REGION Network 39
   RUNG wire#powerrail
      #"8#浊环热水泵引水电磁阀"(READY := wire#w1, HMI_OPEN :=, HMI_CLOSE :=, MA :=, AUTO :=, S :=, JT :=, "TIME" :=, OUT := "8#浊环热水泵引水电磁阀", TIME_OUT =>)
   END_RUNG
   RUNG wire#powerrail
      Contact( "8#浊环热水泵备妥" )
      Contact( "8#浊环热水电动蝶阀备妥" )
   END_RUNG wire#w1
   // the same network as SCL:
   #"8#浊环热水泵引水电磁阀"(READY := "8#浊环热水泵备妥" AND "8#浊环热水电动蝶阀备妥", OUT := "8#浊环热水泵引水电磁阀");   // "引水排气块"
END_REGION

REGION Network 40
   RUNG wire#powerrail
      #"8#浊环热水泵排气电磁阀"(READY := wire#w1, HMI_OPEN :=, HMI_CLOSE :=, MA :=, AUTO :=, S :=, JT :=, "TIME" :=, OUT := "8#浊环热水泵排气电磁阀", TIME_OUT =>)
   END_RUNG
   RUNG wire#powerrail
      Contact( "8#浊环热水泵备妥" )
      Contact( "8#浊环热水电动蝶阀备妥" )
   END_RUNG wire#w1
   // the same network as SCL:
   #"8#浊环热水泵排气电磁阀"(READY := "8#浊环热水泵备妥" AND "8#浊环热水电动蝶阀备妥", OUT := "8#浊环热水泵排气电磁阀");   // "引水排气块"
END_REGION

REGION Network 41
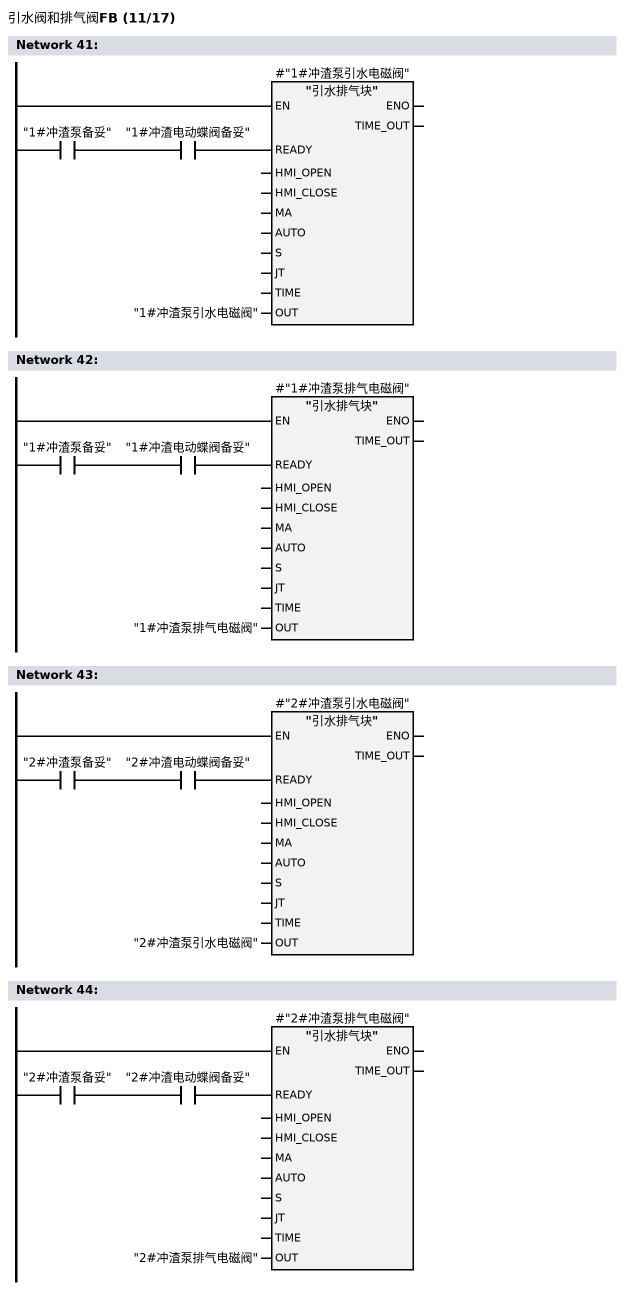
   RUNG wire#powerrail
      #"1#冲渣泵引水电磁阀"(READY := wire#w1, HMI_OPEN :=, HMI_CLOSE :=, MA :=, AUTO :=, S :=, JT :=, "TIME" :=, OUT := "1#冲渣泵引水电磁阀", TIME_OUT =>)
   END_RUNG
   RUNG wire#powerrail
      Contact( "1#冲渣泵备妥" )
      Contact( "1#冲渣电动蝶阀备妥" )
   END_RUNG wire#w1
   // the same network as SCL:
   #"1#冲渣泵引水电磁阀"(READY := "1#冲渣泵备妥" AND "1#冲渣电动蝶阀备妥", OUT := "1#冲渣泵引水电磁阀");   // "引水排气块"
END_REGION

REGION Network 42
   RUNG wire#powerrail
      #"1#冲渣泵排气电磁阀"(READY := wire#w1, HMI_OPEN :=, HMI_CLOSE :=, MA :=, AUTO :=, S :=, JT :=, "TIME" :=, OUT := "1#冲渣泵排气电磁阀", TIME_OUT =>)
   END_RUNG
   RUNG wire#powerrail
      Contact( "1#冲渣泵备妥" )
      Contact( "1#冲渣电动蝶阀备妥" )
   END_RUNG wire#w1
   // the same network as SCL:
   #"1#冲渣泵排气电磁阀"(READY := "1#冲渣泵备妥" AND "1#冲渣电动蝶阀备妥", OUT := "1#冲渣泵排气电磁阀");   // "引水排气块"
END_REGION

REGION Network 43
   RUNG wire#powerrail
      #"2#冲渣泵引水电磁阀"(READY := wire#w1, HMI_OPEN :=, HMI_CLOSE :=, MA :=, AUTO :=, S :=, JT :=, "TIME" :=, OUT := "2#冲渣泵引水电磁阀", TIME_OUT =>)
   END_RUNG
   RUNG wire#powerrail
      Contact( "2#冲渣泵备妥" )
      Contact( "2#冲渣电动蝶阀备妥" )
   END_RUNG wire#w1
   // the same network as SCL:
   #"2#冲渣泵引水电磁阀"(READY := "2#冲渣泵备妥" AND "2#冲渣电动蝶阀备妥", OUT := "2#冲渣泵引水电磁阀");   // "引水排气块"
END_REGION

REGION Network 44
   RUNG wire#powerrail
      #"2#冲渣泵排气电磁阀"(READY := wire#w1, HMI_OPEN :=, HMI_CLOSE :=, MA :=, AUTO :=, S :=, JT :=, "TIME" :=, OUT := "2#冲渣泵排气电磁阀", TIME_OUT =>)
   END_RUNG
   RUNG wire#powerrail
      Contact( "2#冲渣泵备妥" )
      Contact( "2#冲渣电动蝶阀备妥" )
   END_RUNG wire#w1
   // the same network as SCL:
   #"2#冲渣泵排气电磁阀"(READY := "2#冲渣泵备妥" AND "2#冲渣电动蝶阀备妥", OUT := "2#冲渣泵排气电磁阀");   // "引水排气块"
END_REGION

REGION Network 45
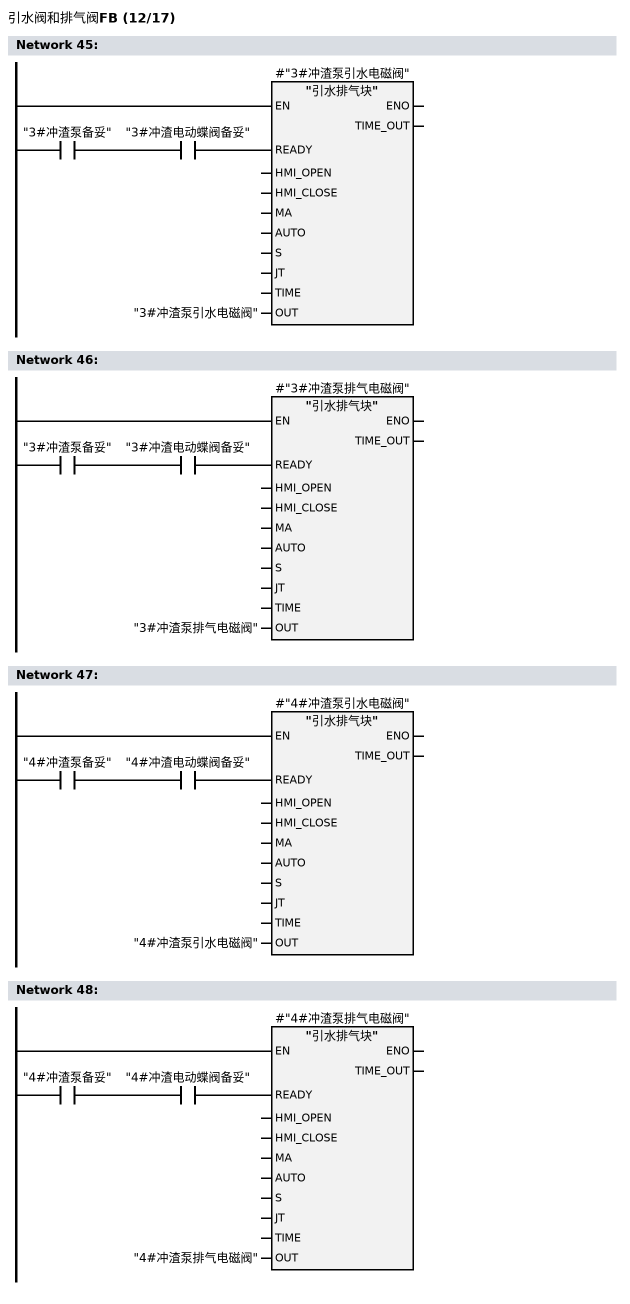
   RUNG wire#powerrail
      #"3#冲渣泵引水电磁阀"(READY := wire#w1, HMI_OPEN :=, HMI_CLOSE :=, MA :=, AUTO :=, S :=, JT :=, "TIME" :=, OUT := "3#冲渣泵引水电磁阀", TIME_OUT =>)
   END_RUNG
   RUNG wire#powerrail
      Contact( "3#冲渣泵备妥" )
      Contact( "3#冲渣电动蝶阀备妥" )
   END_RUNG wire#w1
   // the same network as SCL:
   #"3#冲渣泵引水电磁阀"(READY := "3#冲渣泵备妥" AND "3#冲渣电动蝶阀备妥", OUT := "3#冲渣泵引水电磁阀");   // "引水排气块"
END_REGION

REGION Network 46
   RUNG wire#powerrail
      #"3#冲渣泵排气电磁阀"(READY := wire#w1, HMI_OPEN :=, HMI_CLOSE :=, MA :=, AUTO :=, S :=, JT :=, "TIME" :=, OUT := "3#冲渣泵排气电磁阀", TIME_OUT =>)
   END_RUNG
   RUNG wire#powerrail
      Contact( "3#冲渣泵备妥" )
      Contact( "3#冲渣电动蝶阀备妥" )
   END_RUNG wire#w1
   // the same network as SCL:
   #"3#冲渣泵排气电磁阀"(READY := "3#冲渣泵备妥" AND "3#冲渣电动蝶阀备妥", OUT := "3#冲渣泵排气电磁阀");   // "引水排气块"
END_REGION

REGION Network 47
   RUNG wire#powerrail
      #"4#冲渣泵引水电磁阀"(READY := wire#w1, HMI_OPEN :=, HMI_CLOSE :=, MA :=, AUTO :=, S :=, JT :=, "TIME" :=, OUT := "4#冲渣泵引水电磁阀", TIME_OUT =>)
   END_RUNG
   RUNG wire#powerrail
      Contact( "4#冲渣泵备妥" )
      Contact( "4#冲渣电动蝶阀备妥" )
   END_RUNG wire#w1
   // the same network as SCL:
   #"4#冲渣泵引水电磁阀"(READY := "4#冲渣泵备妥" AND "4#冲渣电动蝶阀备妥", OUT := "4#冲渣泵引水电磁阀");   // "引水排气块"
END_REGION

REGION Network 48
   RUNG wire#powerrail
      #"4#冲渣泵排气电磁阀"(READY := wire#w1, HMI_OPEN :=, HMI_CLOSE :=, MA :=, AUTO :=, S :=, JT :=, "TIME" :=, OUT := "4#冲渣泵排气电磁阀", TIME_OUT =>)
   END_RUNG
   RUNG wire#powerrail
      Contact( "4#冲渣泵备妥" )
      Contact( "4#冲渣电动蝶阀备妥" )
   END_RUNG wire#w1
   // the same network as SCL:
   #"4#冲渣泵排气电磁阀"(READY := "4#冲渣泵备妥" AND "4#冲渣电动蝶阀备妥", OUT := "4#冲渣泵排气电磁阀");   // "引水排气块"
END_REGION

REGION Network 49
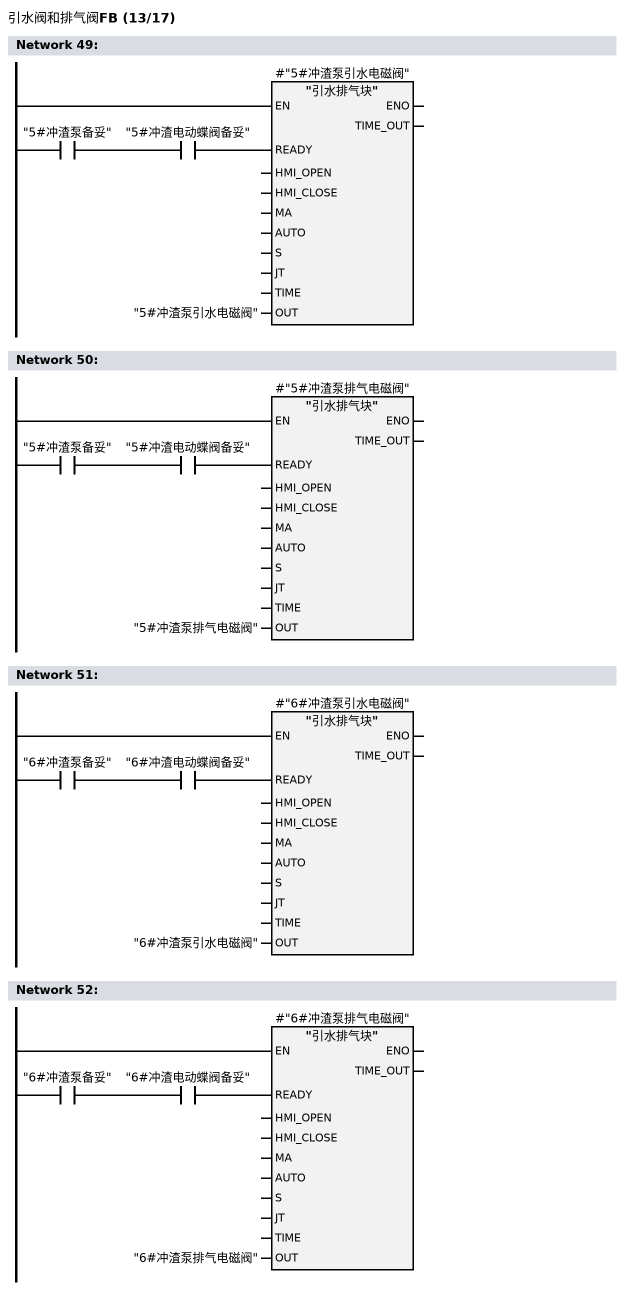
   RUNG wire#powerrail
      #"5#冲渣泵引水电磁阀"(READY := wire#w1, HMI_OPEN :=, HMI_CLOSE :=, MA :=, AUTO :=, S :=, JT :=, "TIME" :=, OUT := "5#冲渣泵引水电磁阀", TIME_OUT =>)
   END_RUNG
   RUNG wire#powerrail
      Contact( "5#冲渣泵备妥" )
      Contact( "5#冲渣电动蝶阀备妥" )
   END_RUNG wire#w1
   // the same network as SCL:
   #"5#冲渣泵引水电磁阀"(READY := "5#冲渣泵备妥" AND "5#冲渣电动蝶阀备妥", OUT := "5#冲渣泵引水电磁阀");   // "引水排气块"
END_REGION

REGION Network 50
   RUNG wire#powerrail
      #"5#冲渣泵排气电磁阀"(READY := wire#w1, HMI_OPEN :=, HMI_CLOSE :=, MA :=, AUTO :=, S :=, JT :=, "TIME" :=, OUT := "5#冲渣泵排气电磁阀", TIME_OUT =>)
   END_RUNG
   RUNG wire#powerrail
      Contact( "5#冲渣泵备妥" )
      Contact( "5#冲渣电动蝶阀备妥" )
   END_RUNG wire#w1
   // the same network as SCL:
   #"5#冲渣泵排气电磁阀"(READY := "5#冲渣泵备妥" AND "5#冲渣电动蝶阀备妥", OUT := "5#冲渣泵排气电磁阀");   // "引水排气块"
END_REGION

REGION Network 51
   RUNG wire#powerrail
      #"6#冲渣泵引水电磁阀"(READY := wire#w1, HMI_OPEN :=, HMI_CLOSE :=, MA :=, AUTO :=, S :=, JT :=, "TIME" :=, OUT := "6#冲渣泵引水电磁阀", TIME_OUT =>)
   END_RUNG
   RUNG wire#powerrail
      Contact( "6#冲渣泵备妥" )
      Contact( "6#冲渣电动蝶阀备妥" )
   END_RUNG wire#w1
   // the same network as SCL:
   #"6#冲渣泵引水电磁阀"(READY := "6#冲渣泵备妥" AND "6#冲渣电动蝶阀备妥", OUT := "6#冲渣泵引水电磁阀");   // "引水排气块"
END_REGION

REGION Network 52
   RUNG wire#powerrail
      #"6#冲渣泵排气电磁阀"(READY := wire#w1, HMI_OPEN :=, HMI_CLOSE :=, MA :=, AUTO :=, S :=, JT :=, "TIME" :=, OUT := "6#冲渣泵排气电磁阀", TIME_OUT =>)
   END_RUNG
   RUNG wire#powerrail
      Contact( "6#冲渣泵备妥" )
      Contact( "6#冲渣电动蝶阀备妥" )
   END_RUNG wire#w1
   // the same network as SCL:
   #"6#冲渣泵排气电磁阀"(READY := "6#冲渣泵备妥" AND "6#冲渣电动蝶阀备妥", OUT := "6#冲渣泵排气电磁阀");   // "引水排气块"
END_REGION

REGION Network 53
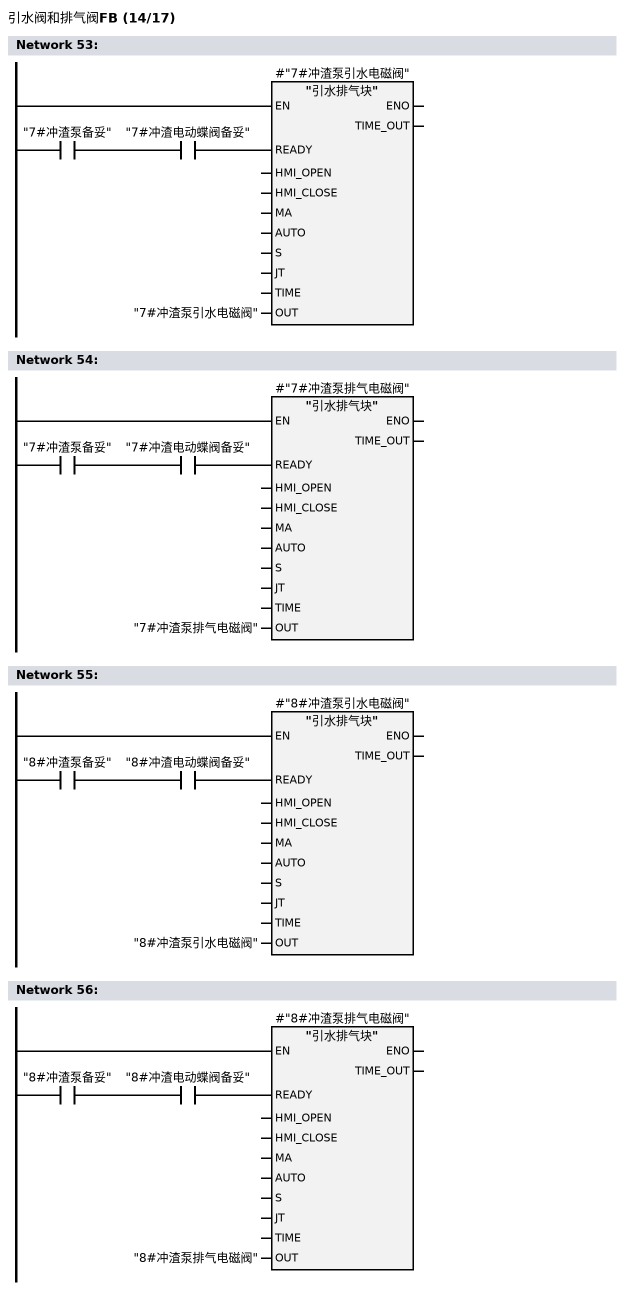
   RUNG wire#powerrail
      #"7#冲渣泵引水电磁阀"(READY := wire#w1, HMI_OPEN :=, HMI_CLOSE :=, MA :=, AUTO :=, S :=, JT :=, "TIME" :=, OUT := "7#冲渣泵引水电磁阀", TIME_OUT =>)
   END_RUNG
   RUNG wire#powerrail
      Contact( "7#冲渣泵备妥" )
      Contact( "7#冲渣电动蝶阀备妥" )
   END_RUNG wire#w1
   // the same network as SCL:
   #"7#冲渣泵引水电磁阀"(READY := "7#冲渣泵备妥" AND "7#冲渣电动蝶阀备妥", OUT := "7#冲渣泵引水电磁阀");   // "引水排气块"
END_REGION

REGION Network 54
   RUNG wire#powerrail
      #"7#冲渣泵排气电磁阀"(READY := wire#w1, HMI_OPEN :=, HMI_CLOSE :=, MA :=, AUTO :=, S :=, JT :=, "TIME" :=, OUT := "7#冲渣泵排气电磁阀", TIME_OUT =>)
   END_RUNG
   RUNG wire#powerrail
      Contact( "7#冲渣泵备妥" )
      Contact( "7#冲渣电动蝶阀备妥" )
   END_RUNG wire#w1
   // the same network as SCL:
   #"7#冲渣泵排气电磁阀"(READY := "7#冲渣泵备妥" AND "7#冲渣电动蝶阀备妥", OUT := "7#冲渣泵排气电磁阀");   // "引水排气块"
END_REGION

REGION Network 55
   RUNG wire#powerrail
      #"8#冲渣泵引水电磁阀"(READY := wire#w1, HMI_OPEN :=, HMI_CLOSE :=, MA :=, AUTO :=, S :=, JT :=, "TIME" :=, OUT := "8#冲渣泵引水电磁阀", TIME_OUT =>)
   END_RUNG
   RUNG wire#powerrail
      Contact( "8#冲渣泵备妥" )
      Contact( "8#冲渣电动蝶阀备妥" )
   END_RUNG wire#w1
   // the same network as SCL:
   #"8#冲渣泵引水电磁阀"(READY := "8#冲渣泵备妥" AND "8#冲渣电动蝶阀备妥", OUT := "8#冲渣泵引水电磁阀");   // "引水排气块"
END_REGION

REGION Network 56
   RUNG wire#powerrail
      #"8#冲渣泵排气电磁阀"(READY := wire#w1, HMI_OPEN :=, HMI_CLOSE :=, MA :=, AUTO :=, S :=, JT :=, "TIME" :=, OUT := "8#冲渣泵排气电磁阀", TIME_OUT =>)
   END_RUNG
   RUNG wire#powerrail
      Contact( "8#冲渣泵备妥" )
      Contact( "8#冲渣电动蝶阀备妥" )
   END_RUNG wire#w1
   // the same network as SCL:
   #"8#冲渣泵排气电磁阀"(READY := "8#冲渣泵备妥" AND "8#冲渣电动蝶阀备妥", OUT := "8#冲渣泵排气电磁阀");   // "引水排气块"
END_REGION

REGION Network 57
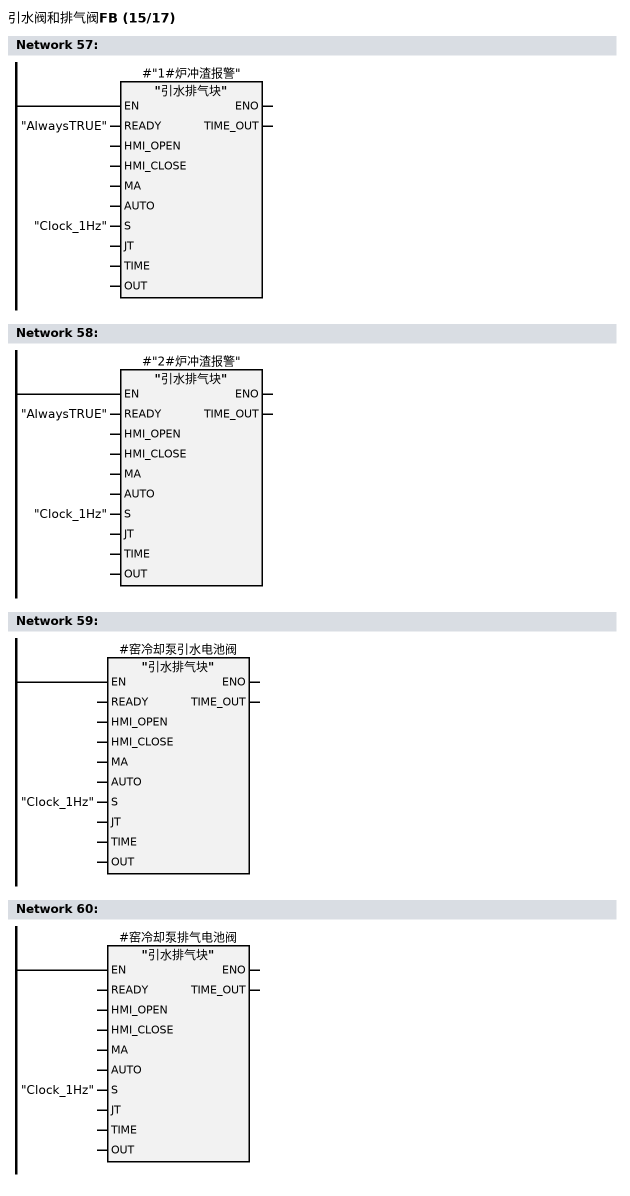
   RUNG wire#powerrail
      #"1#炉冲渣报警"(READY := "AlwaysTRUE", HMI_OPEN :=, HMI_CLOSE :=, MA :=, AUTO :=, S := "Clock_1Hz", JT :=, "TIME" :=, OUT :=, TIME_OUT =>)
   END_RUNG
   // the same network as SCL:
   #"1#炉冲渣报警"(READY := "AlwaysTRUE", S := "Clock_1Hz");   // "引水排气块"
END_REGION

REGION Network 58
   RUNG wire#powerrail
      #"2#炉冲渣报警"(READY := "AlwaysTRUE", HMI_OPEN :=, HMI_CLOSE :=, MA :=, AUTO :=, S := "Clock_1Hz", JT :=, "TIME" :=, OUT :=, TIME_OUT =>)
   END_RUNG
   // the same network as SCL:
   #"2#炉冲渣报警"(READY := "AlwaysTRUE", S := "Clock_1Hz");   // "引水排气块"
END_REGION

REGION Network 59
   RUNG wire#powerrail
      #窑冷却泵引水电池阀(READY :=, HMI_OPEN :=, HMI_CLOSE :=, MA :=, AUTO :=, S := "Clock_1Hz", JT :=, "TIME" :=, OUT :=, TIME_OUT =>)
   END_RUNG
   // the same network as SCL:
   #窑冷却泵引水电池阀(S := "Clock_1Hz");   // "引水排气块"
END_REGION

REGION Network 60
   RUNG wire#powerrail
      #窑冷却泵排气电池阀(READY :=, HMI_OPEN :=, HMI_CLOSE :=, MA :=, AUTO :=, S := "Clock_1Hz", JT :=, "TIME" :=, OUT :=, TIME_OUT =>)
   END_RUNG
   // the same network as SCL:
   #窑冷却泵排气电池阀(S := "Clock_1Hz");   // "引水排气块"
END_REGION

REGION Network 61
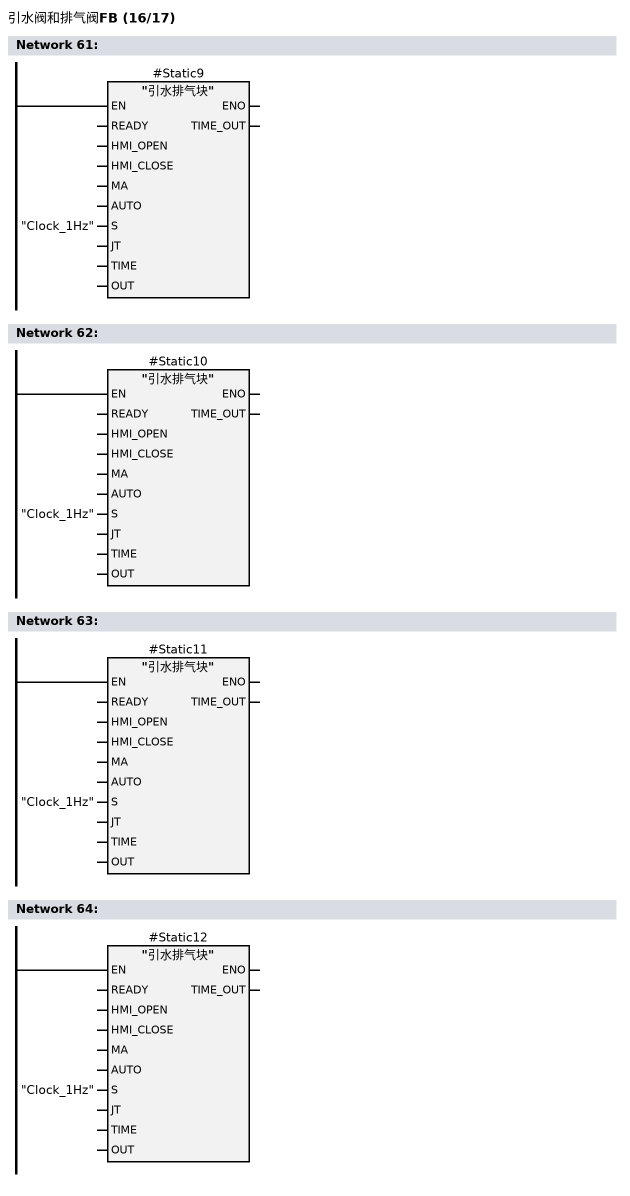
   RUNG wire#powerrail
      #Static9(READY :=, HMI_OPEN :=, HMI_CLOSE :=, MA :=, AUTO :=, S := "Clock_1Hz", JT :=, "TIME" :=, OUT :=, TIME_OUT =>)
   END_RUNG
   // the same network as SCL:
   #Static9(S := "Clock_1Hz");   // "引水排气块"
END_REGION

REGION Network 62
   RUNG wire#powerrail
      #Static10(READY :=, HMI_OPEN :=, HMI_CLOSE :=, MA :=, AUTO :=, S := "Clock_1Hz", JT :=, "TIME" :=, OUT :=, TIME_OUT =>)
   END_RUNG
   // the same network as SCL:
   #Static10(S := "Clock_1Hz");   // "引水排气块"
END_REGION

REGION Network 63
   RUNG wire#powerrail
      #Static11(READY :=, HMI_OPEN :=, HMI_CLOSE :=, MA :=, AUTO :=, S := "Clock_1Hz", JT :=, "TIME" :=, OUT :=, TIME_OUT =>)
   END_RUNG
   // the same network as SCL:
   #Static11(S := "Clock_1Hz");   // "引水排气块"
END_REGION

REGION Network 64
   RUNG wire#powerrail
      #Static12(READY :=, HMI_OPEN :=, HMI_CLOSE :=, MA :=, AUTO :=, S := "Clock_1Hz", JT :=, "TIME" :=, OUT :=, TIME_OUT =>)
   END_RUNG
   // the same network as SCL:
   #Static12(S := "Clock_1Hz");   // "引水排气块"
END_REGION

REGION Network 65
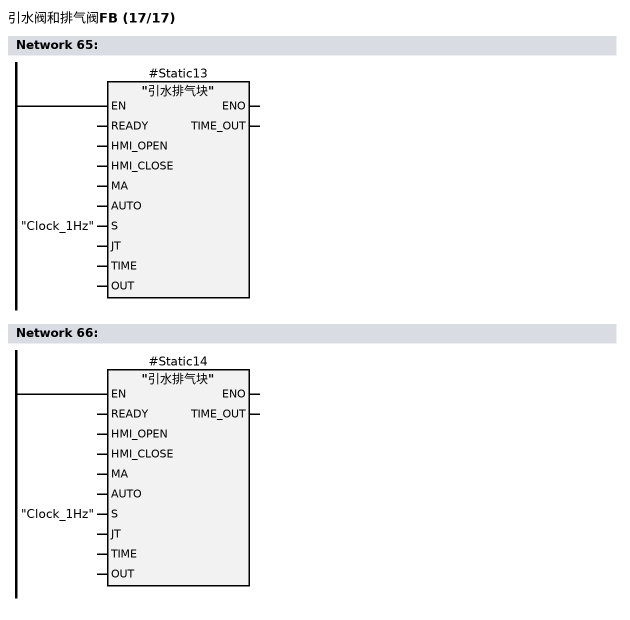
   RUNG wire#powerrail
      #Static13(READY :=, HMI_OPEN :=, HMI_CLOSE :=, MA :=, AUTO :=, S := "Clock_1Hz", JT :=, "TIME" :=, OUT :=, TIME_OUT =>)
   END_RUNG
   // the same network as SCL:
   #Static13(S := "Clock_1Hz");   // "引水排气块"
END_REGION

REGION Network 66
   RUNG wire#powerrail
      #Static14(READY :=, HMI_OPEN :=, HMI_CLOSE :=, MA :=, AUTO :=, S := "Clock_1Hz", JT :=, "TIME" :=, OUT :=, TIME_OUT =>)
   END_RUNG
   // the same network as SCL:
   #Static14(S := "Clock_1Hz");   // "引水排气块"
END_REGION
END_FUNCTION_BLOCK

FUNCTION_BLOCK "电机_泵FB"   // FB13, LAD
{ S7_Optimized_Access := 'FALSE' }
VERSION : 0.1
   VAR
      "1#冲渣泵驱动" : "电机_冷却塔风机";
      "2#冲渣泵驱动" : "电机_冷却塔风机";
      "3#冲渣泵驱动" : "电机_冷却塔风机";
      "4#冲渣泵驱动" : "电机_冷却塔风机";
      "5#冲渣泵驱动" : "电机_冷却塔风机";
      "6#冲渣泵驱动" : "电机_冷却塔风机";
      "7#冲渣泵驱动" : "电机_冷却塔风机";
      "8#冲渣泵驱动" : "电机_冷却塔风机";
      "1#浊环热水泵驱动" : "电机_冷却塔风机";
      "2#浊环热水泵驱动" : "电机_冷却塔风机";
      "3#浊环热水泵驱动" : "电机_冷却塔风机";
      "4#浊环热水泵驱动" : "电机_冷却塔风机";
      "5#浊环热水泵驱动" : "电机_冷却塔风机";
      "6#浊环热水泵驱动" : "电机_冷却塔风机";
      "7#浊环热水泵驱动" : "电机_冷却塔风机";
      "8#浊环热水泵驱动" : "电机_冷却塔风机";
      "1#炉体循环水泵驱动" : "电机_冷却塔风机";
      "2#炉体循环水泵驱动" : "电机_冷却塔风机";
      "3#炉体循环水泵驱动" : "电机_冷却塔风机";
      "1#电极循环水泵驱动" : "电机_冷却塔风机";
      "2#电极循环水泵驱动" : "电机_冷却塔风机";
      "3#电极循环水泵驱动" : "电机_冷却塔风机";
      "4#电极循环水泵驱动" : "电机_冷却塔风机";
      "1#净环热水泵驱动" : "电机_冷却塔风机";
      "2#净环热水泵驱动" : "电机_冷却塔风机";
      "3#净环热水泵驱动" : "电机_冷却塔风机";
      "4#净环热水泵驱动" : "电机_冷却塔风机";
      "5#净环热水泵驱动" : "电机_冷却塔风机";
      "1#柴油泵驱动" : "电机_冷却塔风机";
      "2#柴油泵驱动" : "电机_冷却塔风机";
      窑冷却泵驱动 : "电机_冷却塔风机";
      Static1 : "电机_冷却塔风机";
      Static2 : "电机_冷却塔风机";
      Static3 : "电机_冷却塔风机";
      Static4 : "电机_冷却塔风机";
      Static5 : "电机_冷却塔风机";
      Static6 : "电机_冷却塔风机";
      Static7 : "电机_冷却塔风机";
      Static8 : "电机_冷却塔风机";
      Static9 : "电机_冷却塔风机";
      Static10 : "电机_冷却塔风机";
      Static11 : "电机_冷却塔风机";
      Static12 : "电机_冷却塔风机";
      Static13 : "电机_冷却塔风机";
      Static14 : "电机_冷却塔风机";
      Static15 : "电机_冷却塔风机";
      Static16 : "电机_冷却塔风机";
      Static17 : "电机_冷却塔风机";
      Static18 : "电机_冷却塔风机";
      Static19 : "电机_冷却塔风机";
      Static20 : "电机_冷却塔风机";
      Static21 : "电机_冷却塔风机";
      Static22 : "电机_冷却塔风机";
      Static23 : "电机_冷却塔风机";
      Static24 : "电机_冷却塔风机";
      Static25 : "电机_冷却塔风机";
      Static26 : "电机_冷却塔风机";
      Static27 : "电机_冷却塔风机";
      Static28 : "电机_冷却塔风机";
      Static29 : "电机_冷却塔风机";
      Static30 : "电机_冷却塔风机";
      Static31 : "电机_冷却塔风机";
      Static32 : "电机_冷却塔风机";
      Static33 : "电机_冷却塔风机";
      Static34 : "电机_冷却塔风机";
      Static35 : "电机_冷却塔风机";
      Static36 : "电机_冷却塔风机";
      Static37 : "电机_冷却塔风机";
      Static38 : "电机_冷却塔风机";
      Static39 : "电机_冷却塔风机";
      Static40 : "电机_冷却塔风机";
      Static41 : "电机_冷却塔风机";
      Static42 : "电机_冷却塔风机";
      Static43 : "电机_冷却塔风机";
      Static44 : "电机_冷却塔风机";
      Static45 : "电机_冷却塔风机";
      Static46 : "电机_冷却塔风机";
      Static47 : "电机_冷却塔风机";
      Static48 : "电机_冷却塔风机";
      Static49 : "电机_冷却塔风机";
   END_VAR
BEGIN

REGION Network 1
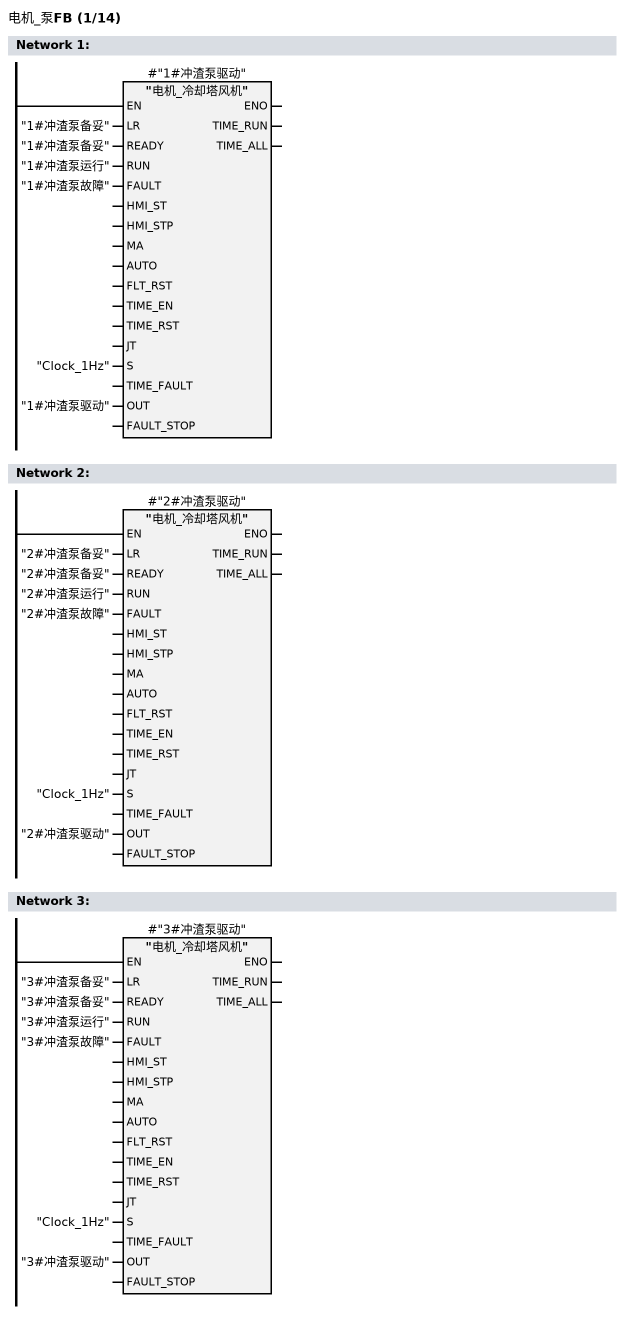
   RUNG wire#powerrail
      #"1#冲渣泵驱动"(LR := "1#冲渣泵备妥", READY := "1#冲渣泵备妥", RUN := "1#冲渣泵运行", FAULT := "1#冲渣泵故障", HMI_ST :=, HMI_STP :=, MA :=, AUTO :=, FLT_RST :=, TIME_EN :=, TIME_RST :=, JT :=, S := "Clock_1Hz", TIME_FAULT :=, OUT := "1#冲渣泵驱动", FAULT_STOP :=, TIME_RUN =>, TIME_ALL =>)
   END_RUNG
   // the same network as SCL:
   #"1#冲渣泵驱动"(LR := "1#冲渣泵备妥",   // "电机_冷却塔风机"
              READY := "1#冲渣泵备妥",
              RUN := "1#冲渣泵运行",
              FAULT := "1#冲渣泵故障",
              S := "Clock_1Hz",
              OUT := "1#冲渣泵驱动");
END_REGION

REGION Network 2
   RUNG wire#powerrail
      #"2#冲渣泵驱动"(LR := "2#冲渣泵备妥", READY := "2#冲渣泵备妥", RUN := "2#冲渣泵运行", FAULT := "2#冲渣泵故障", HMI_ST :=, HMI_STP :=, MA :=, AUTO :=, FLT_RST :=, TIME_EN :=, TIME_RST :=, JT :=, S := "Clock_1Hz", TIME_FAULT :=, OUT := "2#冲渣泵驱动", FAULT_STOP :=, TIME_RUN =>, TIME_ALL =>)
   END_RUNG
   // the same network as SCL:
   #"2#冲渣泵驱动"(LR := "2#冲渣泵备妥",   // "电机_冷却塔风机"
              READY := "2#冲渣泵备妥",
              RUN := "2#冲渣泵运行",
              FAULT := "2#冲渣泵故障",
              S := "Clock_1Hz",
              OUT := "2#冲渣泵驱动");
END_REGION

REGION Network 3
   RUNG wire#powerrail
      #"3#冲渣泵驱动"(LR := "3#冲渣泵备妥", READY := "3#冲渣泵备妥", RUN := "3#冲渣泵运行", FAULT := "3#冲渣泵故障", HMI_ST :=, HMI_STP :=, MA :=, AUTO :=, FLT_RST :=, TIME_EN :=, TIME_RST :=, JT :=, S := "Clock_1Hz", TIME_FAULT :=, OUT := "3#冲渣泵驱动", FAULT_STOP :=, TIME_RUN =>, TIME_ALL =>)
   END_RUNG
   // the same network as SCL:
   #"3#冲渣泵驱动"(LR := "3#冲渣泵备妥",   // "电机_冷却塔风机"
              READY := "3#冲渣泵备妥",
              RUN := "3#冲渣泵运行",
              FAULT := "3#冲渣泵故障",
              S := "Clock_1Hz",
              OUT := "3#冲渣泵驱动");
END_REGION

REGION Network 4
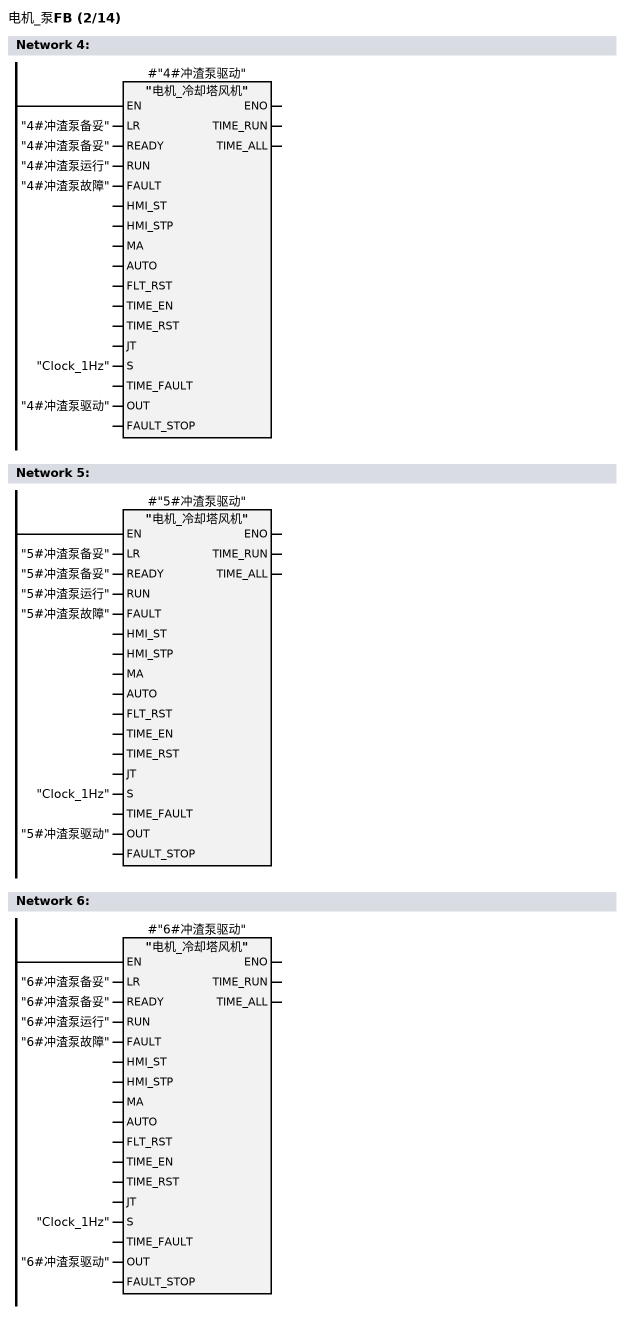
   RUNG wire#powerrail
      #"4#冲渣泵驱动"(LR := "4#冲渣泵备妥", READY := "4#冲渣泵备妥", RUN := "4#冲渣泵运行", FAULT := "4#冲渣泵故障", HMI_ST :=, HMI_STP :=, MA :=, AUTO :=, FLT_RST :=, TIME_EN :=, TIME_RST :=, JT :=, S := "Clock_1Hz", TIME_FAULT :=, OUT := "4#冲渣泵驱动", FAULT_STOP :=, TIME_RUN =>, TIME_ALL =>)
   END_RUNG
   // the same network as SCL:
   #"4#冲渣泵驱动"(LR := "4#冲渣泵备妥",   // "电机_冷却塔风机"
              READY := "4#冲渣泵备妥",
              RUN := "4#冲渣泵运行",
              FAULT := "4#冲渣泵故障",
              S := "Clock_1Hz",
              OUT := "4#冲渣泵驱动");
END_REGION

REGION Network 5
   RUNG wire#powerrail
      #"5#冲渣泵驱动"(LR := "5#冲渣泵备妥", READY := "5#冲渣泵备妥", RUN := "5#冲渣泵运行", FAULT := "5#冲渣泵故障", HMI_ST :=, HMI_STP :=, MA :=, AUTO :=, FLT_RST :=, TIME_EN :=, TIME_RST :=, JT :=, S := "Clock_1Hz", TIME_FAULT :=, OUT := "5#冲渣泵驱动", FAULT_STOP :=, TIME_RUN =>, TIME_ALL =>)
   END_RUNG
   // the same network as SCL:
   #"5#冲渣泵驱动"(LR := "5#冲渣泵备妥",   // "电机_冷却塔风机"
              READY := "5#冲渣泵备妥",
              RUN := "5#冲渣泵运行",
              FAULT := "5#冲渣泵故障",
              S := "Clock_1Hz",
              OUT := "5#冲渣泵驱动");
END_REGION

REGION Network 6
   RUNG wire#powerrail
      #"6#冲渣泵驱动"(LR := "6#冲渣泵备妥", READY := "6#冲渣泵备妥", RUN := "6#冲渣泵运行", FAULT := "6#冲渣泵故障", HMI_ST :=, HMI_STP :=, MA :=, AUTO :=, FLT_RST :=, TIME_EN :=, TIME_RST :=, JT :=, S := "Clock_1Hz", TIME_FAULT :=, OUT := "6#冲渣泵驱动", FAULT_STOP :=, TIME_RUN =>, TIME_ALL =>)
   END_RUNG
   // the same network as SCL:
   #"6#冲渣泵驱动"(LR := "6#冲渣泵备妥",   // "电机_冷却塔风机"
              READY := "6#冲渣泵备妥",
              RUN := "6#冲渣泵运行",
              FAULT := "6#冲渣泵故障",
              S := "Clock_1Hz",
              OUT := "6#冲渣泵驱动");
END_REGION

REGION Network 7
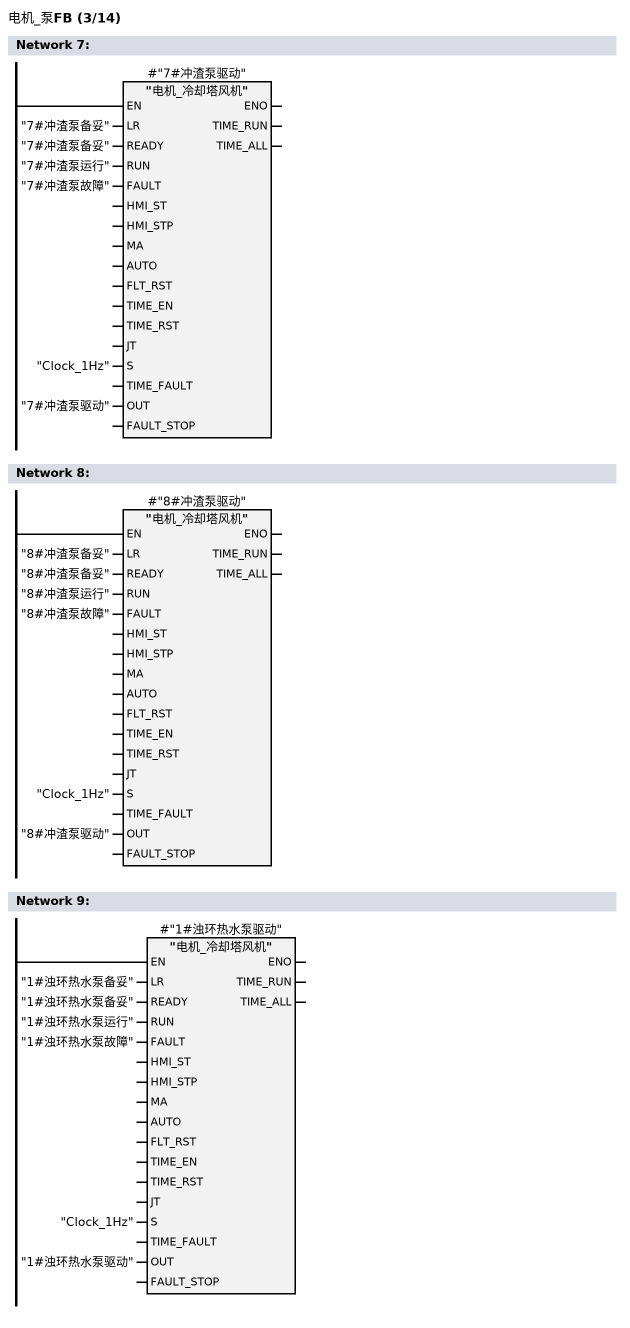
   RUNG wire#powerrail
      #"7#冲渣泵驱动"(LR := "7#冲渣泵备妥", READY := "7#冲渣泵备妥", RUN := "7#冲渣泵运行", FAULT := "7#冲渣泵故障", HMI_ST :=, HMI_STP :=, MA :=, AUTO :=, FLT_RST :=, TIME_EN :=, TIME_RST :=, JT :=, S := "Clock_1Hz", TIME_FAULT :=, OUT := "7#冲渣泵驱动", FAULT_STOP :=, TIME_RUN =>, TIME_ALL =>)
   END_RUNG
   // the same network as SCL:
   #"7#冲渣泵驱动"(LR := "7#冲渣泵备妥",   // "电机_冷却塔风机"
              READY := "7#冲渣泵备妥",
              RUN := "7#冲渣泵运行",
              FAULT := "7#冲渣泵故障",
              S := "Clock_1Hz",
              OUT := "7#冲渣泵驱动");
END_REGION

REGION Network 8
   RUNG wire#powerrail
      #"8#冲渣泵驱动"(LR := "8#冲渣泵备妥", READY := "8#冲渣泵备妥", RUN := "8#冲渣泵运行", FAULT := "8#冲渣泵故障", HMI_ST :=, HMI_STP :=, MA :=, AUTO :=, FLT_RST :=, TIME_EN :=, TIME_RST :=, JT :=, S := "Clock_1Hz", TIME_FAULT :=, OUT := "8#冲渣泵驱动", FAULT_STOP :=, TIME_RUN =>, TIME_ALL =>)
   END_RUNG
   // the same network as SCL:
   #"8#冲渣泵驱动"(LR := "8#冲渣泵备妥",   // "电机_冷却塔风机"
              READY := "8#冲渣泵备妥",
              RUN := "8#冲渣泵运行",
              FAULT := "8#冲渣泵故障",
              S := "Clock_1Hz",
              OUT := "8#冲渣泵驱动");
END_REGION

REGION Network 9
   RUNG wire#powerrail
      #"1#浊环热水泵驱动"(LR := "1#浊环热水泵备妥", READY := "1#浊环热水泵备妥", RUN := "1#浊环热水泵运行", FAULT := "1#浊环热水泵故障", HMI_ST :=, HMI_STP :=, MA :=, AUTO :=, FLT_RST :=, TIME_EN :=, TIME_RST :=, JT :=, S := "Clock_1Hz", TIME_FAULT :=, OUT := "1#浊环热水泵驱动", FAULT_STOP :=, TIME_RUN =>, TIME_ALL =>)
   END_RUNG
   // the same network as SCL:
   #"1#浊环热水泵驱动"(LR := "1#浊环热水泵备妥",   // "电机_冷却塔风机"
                READY := "1#浊环热水泵备妥",
                RUN := "1#浊环热水泵运行",
                FAULT := "1#浊环热水泵故障",
                S := "Clock_1Hz",
                OUT := "1#浊环热水泵驱动");
END_REGION

REGION Network 10
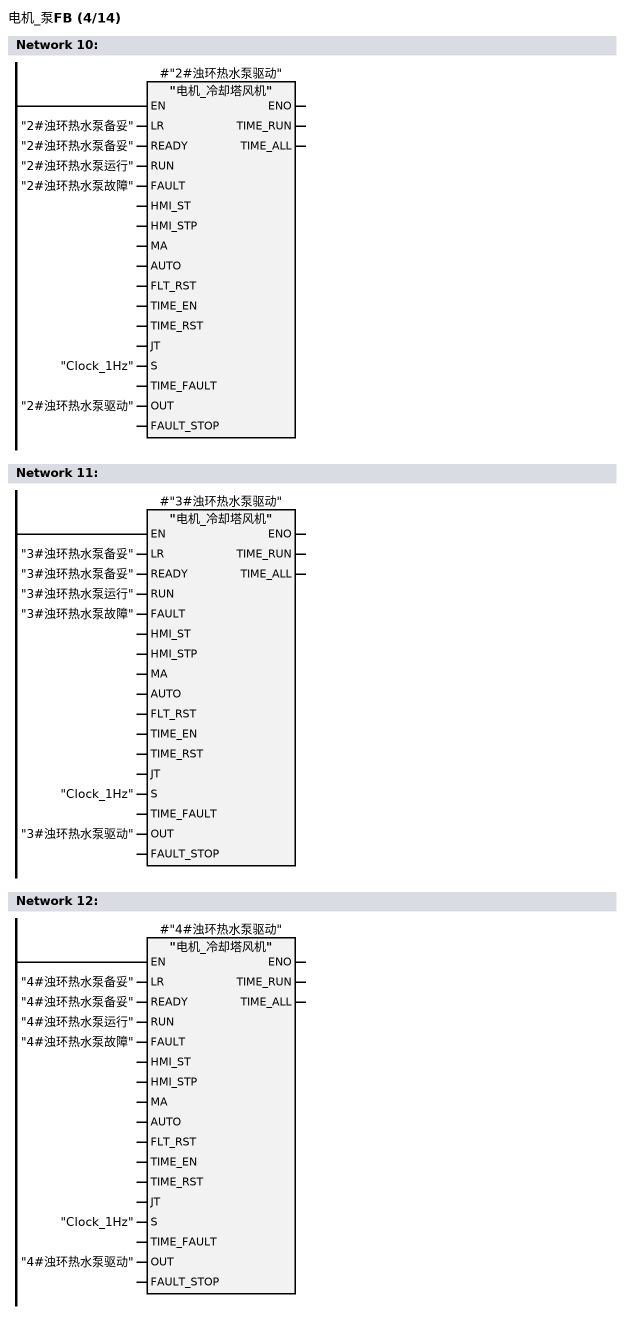
   RUNG wire#powerrail
      #"2#浊环热水泵驱动"(LR := "2#浊环热水泵备妥", READY := "2#浊环热水泵备妥", RUN := "2#浊环热水泵运行", FAULT := "2#浊环热水泵故障", HMI_ST :=, HMI_STP :=, MA :=, AUTO :=, FLT_RST :=, TIME_EN :=, TIME_RST :=, JT :=, S := "Clock_1Hz", TIME_FAULT :=, OUT := "2#浊环热水泵驱动", FAULT_STOP :=, TIME_RUN =>, TIME_ALL =>)
   END_RUNG
   // the same network as SCL:
   #"2#浊环热水泵驱动"(LR := "2#浊环热水泵备妥",   // "电机_冷却塔风机"
                READY := "2#浊环热水泵备妥",
                RUN := "2#浊环热水泵运行",
                FAULT := "2#浊环热水泵故障",
                S := "Clock_1Hz",
                OUT := "2#浊环热水泵驱动");
END_REGION

REGION Network 11
   RUNG wire#powerrail
      #"3#浊环热水泵驱动"(LR := "3#浊环热水泵备妥", READY := "3#浊环热水泵备妥", RUN := "3#浊环热水泵运行", FAULT := "3#浊环热水泵故障", HMI_ST :=, HMI_STP :=, MA :=, AUTO :=, FLT_RST :=, TIME_EN :=, TIME_RST :=, JT :=, S := "Clock_1Hz", TIME_FAULT :=, OUT := "3#浊环热水泵驱动", FAULT_STOP :=, TIME_RUN =>, TIME_ALL =>)
   END_RUNG
   // the same network as SCL:
   #"3#浊环热水泵驱动"(LR := "3#浊环热水泵备妥",   // "电机_冷却塔风机"
                READY := "3#浊环热水泵备妥",
                RUN := "3#浊环热水泵运行",
                FAULT := "3#浊环热水泵故障",
                S := "Clock_1Hz",
                OUT := "3#浊环热水泵驱动");
END_REGION

REGION Network 12
   RUNG wire#powerrail
      #"4#浊环热水泵驱动"(LR := "4#浊环热水泵备妥", READY := "4#浊环热水泵备妥", RUN := "4#浊环热水泵运行", FAULT := "4#浊环热水泵故障", HMI_ST :=, HMI_STP :=, MA :=, AUTO :=, FLT_RST :=, TIME_EN :=, TIME_RST :=, JT :=, S := "Clock_1Hz", TIME_FAULT :=, OUT := "4#浊环热水泵驱动", FAULT_STOP :=, TIME_RUN =>, TIME_ALL =>)
   END_RUNG
   // the same network as SCL:
   #"4#浊环热水泵驱动"(LR := "4#浊环热水泵备妥",   // "电机_冷却塔风机"
                READY := "4#浊环热水泵备妥",
                RUN := "4#浊环热水泵运行",
                FAULT := "4#浊环热水泵故障",
                S := "Clock_1Hz",
                OUT := "4#浊环热水泵驱动");
END_REGION

REGION Network 13
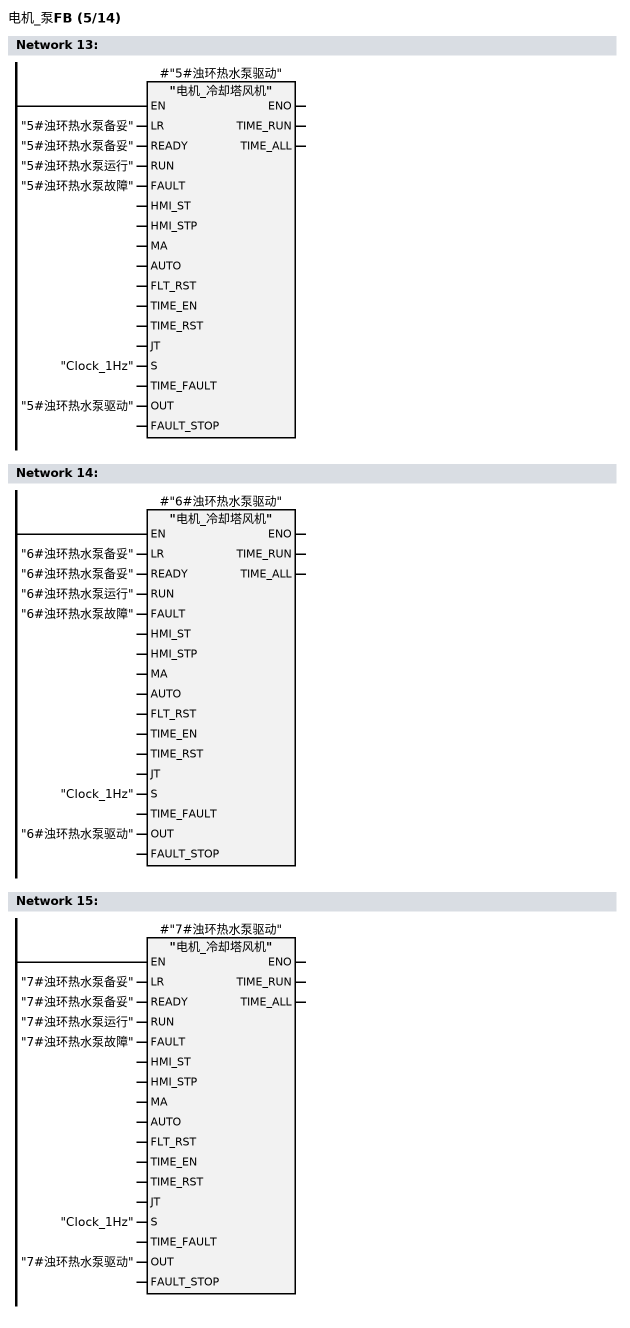
   RUNG wire#powerrail
      #"5#浊环热水泵驱动"(LR := "5#浊环热水泵备妥", READY := "5#浊环热水泵备妥", RUN := "5#浊环热水泵运行", FAULT := "5#浊环热水泵故障", HMI_ST :=, HMI_STP :=, MA :=, AUTO :=, FLT_RST :=, TIME_EN :=, TIME_RST :=, JT :=, S := "Clock_1Hz", TIME_FAULT :=, OUT := "5#浊环热水泵驱动", FAULT_STOP :=, TIME_RUN =>, TIME_ALL =>)
   END_RUNG
   // the same network as SCL:
   #"5#浊环热水泵驱动"(LR := "5#浊环热水泵备妥",   // "电机_冷却塔风机"
                READY := "5#浊环热水泵备妥",
                RUN := "5#浊环热水泵运行",
                FAULT := "5#浊环热水泵故障",
                S := "Clock_1Hz",
                OUT := "5#浊环热水泵驱动");
END_REGION

REGION Network 14
   RUNG wire#powerrail
      #"6#浊环热水泵驱动"(LR := "6#浊环热水泵备妥", READY := "6#浊环热水泵备妥", RUN := "6#浊环热水泵运行", FAULT := "6#浊环热水泵故障", HMI_ST :=, HMI_STP :=, MA :=, AUTO :=, FLT_RST :=, TIME_EN :=, TIME_RST :=, JT :=, S := "Clock_1Hz", TIME_FAULT :=, OUT := "6#浊环热水泵驱动", FAULT_STOP :=, TIME_RUN =>, TIME_ALL =>)
   END_RUNG
   // the same network as SCL:
   #"6#浊环热水泵驱动"(LR := "6#浊环热水泵备妥",   // "电机_冷却塔风机"
                READY := "6#浊环热水泵备妥",
                RUN := "6#浊环热水泵运行",
                FAULT := "6#浊环热水泵故障",
                S := "Clock_1Hz",
                OUT := "6#浊环热水泵驱动");
END_REGION

REGION Network 15
   RUNG wire#powerrail
      #"7#浊环热水泵驱动"(LR := "7#浊环热水泵备妥", READY := "7#浊环热水泵备妥", RUN := "7#浊环热水泵运行", FAULT := "7#浊环热水泵故障", HMI_ST :=, HMI_STP :=, MA :=, AUTO :=, FLT_RST :=, TIME_EN :=, TIME_RST :=, JT :=, S := "Clock_1Hz", TIME_FAULT :=, OUT := "7#浊环热水泵驱动", FAULT_STOP :=, TIME_RUN =>, TIME_ALL =>)
   END_RUNG
   // the same network as SCL:
   #"7#浊环热水泵驱动"(LR := "7#浊环热水泵备妥",   // "电机_冷却塔风机"
                READY := "7#浊环热水泵备妥",
                RUN := "7#浊环热水泵运行",
                FAULT := "7#浊环热水泵故障",
                S := "Clock_1Hz",
                OUT := "7#浊环热水泵驱动");
END_REGION

REGION Network 16
